FUNCTION "Get Station Selection Number" : Void   // FC16, SCL
{ S7_Optimized_Access := 'TRUE' }
VERSION : 0.1
   VAR_INPUT
      next : Bool;   // 'next' or 'prev'
      prev : Bool;
      stations : "Stations";
   END_VAR
   VAR_IN_OUT
      selStnNumber : Int;
   END_VAR
   VAR_TEMP
      i : Int;
      stnCount : Int;
      stnSelected : Bool;
   END_VAR
BEGIN
   REGION "COPY TO LOCAL"
       #stnCount := "stnCount";
   END_REGION

   REGION "INITIALIZE INDEX"
       #i := #selStnNumber;
   END_REGION

   REGION "PREVIOUS MODE"

       REGION "DECREMENT"
           IF #prev THEN
               #i -= 1;
           END_IF;
       END_REGION

       REGION "LOW LIMIT ROLLOVER"
           IF #i < 0 THEN
               #i := #stnCount;
           END_IF;
       END_REGION

   END_REGION

   REGION "NEXT MODE"

       REGION "INCREMENT"
           IF #next THEN
               #i += 1;
           END_IF;
       END_REGION

       REGION "HIGH LIMIT ROLLOVER"
           IF #i > #stnCount THEN
               #i := 0;
           END_IF;
       END_REGION

   END_REGION

   REGION "COPY TO LOCAL"
       #stnSelected := #stations.me[#i].settings.selected;
   END_REGION

   REGION "FIND NEXT SELECTED STATION"
       WHILE NOT #stnSelected DO

           REGION "PREVIOUS MODE"

               REGION "DECREMENT"
                   IF #prev THEN
                       #i -= 1;
                   END_IF;
               END_REGION

               REGION "LOW LIMIT ROLLOVER"
                   IF #i < 0 THEN
                       #i := #stnCount;
                   END_IF;
               END_REGION

           END_REGION

           REGION "NEXT MODE"

               REGION "INCREMENT"
                   IF #next THEN
                       #i += 1;
                   END_IF;
               END_REGION

               REGION "HIGH LIMIT ROLLOVER"
                   IF #i > #stnCount THEN
                       #i := 0;
                   END_IF;
               END_REGION

           END_REGION

           REGION "SAVE WHILE CONDITION"
               #stnSelected := #stations.me[#i].settings.selected;
           END_REGION

       END_WHILE;
   END_REGION

   REGION "RETURN VALUE"
       #selStnNumber := #i;
   END_REGION
END_FUNCTION

FUNCTION "Populate Button Details" : Void   // FC17, SCL
{ S7_Optimized_Access := 'TRUE' }
VERSION : 0.1
   VAR_INPUT
      selStnNumber : Int;
      stations : "Stations";
   END_VAR
   VAR_IN_OUT
      settings : "Settings";
   END_VAR
   VAR_TEMP
      btnCount : Int;
      i : Int;
      partNumber : WString;
      pBtn : Int;
      timerWS : WString;
   END_VAR
BEGIN
   REGION "COPY TO LOCAL"
       #btnCount := "ptsPerStn";
   END_REGION

   REGION "FOR EACH BUTTON"
       FOR #i := 0 TO #btnCount DO

           REGION "CALCULATE BUTTON POINTER"
               IF #i MOD 2 = 0 THEN
                   #pBtn := 7 - #i / 2;
               END_IF;
               IF #i MOD 2 <> 0 THEN
                   #pBtn := 3 - #i / 2;
               END_IF;
           END_REGION

           REGION "BUTTON LABEL"
               #settings.viewingStation.btns[#i].label.value := "Strip Sign"(INT_TO_WSTRING(#i + 1));
           END_REGION

           REGION "ALLOTTED TIME"
               #timerWS := "Real to WString Timer"(#stations.me[#selStnNumber].presetTime.allotted[#pBtn]);
               #settings.viewingStation.btns[#i].alloted.value := #timerWS;
           END_REGION

           REGION "CRITICAL TIME"
               #timerWS := "Real to WString Timer"(#stations.me[#selStnNumber].presetTime.critical[#pBtn]);
               #settings.viewingStation.btns[#i].critical.value := #timerWS;
           END_REGION

           REGION "PART NUMBER"
               #partNumber := #stations.me[#selStnNumber].partNumbers[#pBtn];
               #settings.viewingStation.btns[#i].partNumber.value := #partNumber;
           END_REGION

       END_FOR;
   END_REGION
END_FUNCTION

FUNCTION "Assign Station Parameters" : Void   // FC18, SCL
{ S7_Optimized_Access := 'TRUE' }
VERSION : 0.1
   VAR_IN_OUT
      settings : "Settings";
      stations : "Stations";
   END_VAR
   VAR_TEMP
      dzEntered : Bool;
      dzLabel : WString;
      i : Int;
      lineEntered : Bool;
      lineLabel : WString;
      stnCount : Int;
      stnSelected : Bool;
   END_VAR
BEGIN
   REGION "COPY TO LOCAL"    
       #dzEntered := #settings.viewingStation.dzData.inputFinished;
       #lineEntered := #settings.viewingStation.lineData.inputFinished;
       #stnCount := "stnCount";
   END_REGION

   REGION "ON PARAMETER ENTRY"
       IF #dzEntered OR #lineEntered THEN

           REGION "TURN OFF THE LIGHTS"
               #settings.viewingStation.dzData.inputFinished := FALSE;
               #settings.viewingStation.lineData.inputFinished := FALSE;
           END_REGION

           REGION "FOR EACH STATION"
               FOR #i := 0 TO #stnCount DO

                   REGION "COPY TO LOCAL"
                       #stnSelected := #stations.me[#i].settings.selected;
                   END_REGION

                   REGION "ON SELECTED STATION"
                       IF #stnSelected THEN

                           REGION "ON DROP ZONE INPUT"
                               IF #dzEntered THEN

                                   REGION "GET FROM HMI"
                                       #dzLabel := #settings.viewingStation.dzData.value;
                                   END_REGION

                                   REGION "WRITE TO STATION PARAMETER"
                                       #stations.me[#i].dropZone := WSTRING_TO_USINT(#dzLabel);
                                   END_REGION

                               END_IF;
                           END_REGION

                           REGION "ON LINE LABEL INPUT"
                               IF #lineEntered THEN

                                   REGION "GET FROM HMI"
                                       #lineLabel := #settings.viewingStation.lineData.value;
                                   END_REGION

                                   REGION "WRITE TO STATION PARAMETER"
                                       #stations.me[#i].line := #lineLabel;
                                   END_REGION

                               END_IF;
                           END_REGION

                       END_IF;
                   END_REGION

               END_FOR;
           END_REGION

       END_IF;
   END_REGION
END_FUNCTION

FUNCTION "Animate Button Details" : Void   // FC19, SCL
{ S7_Optimized_Access := 'TRUE' }
VERSION : 0.1
   VAR_INPUT
      stations : "Stations";
   END_VAR
   VAR_IN_OUT
      settings : "Settings";
   END_VAR
   VAR_TEMP
      animate : USInt;
      btnCount : Int;
      btnSelected : Bool;
      deselected : USInt;
      i : Int;
      invisible : USInt;
      pBtn : Int;
      selected : USInt;
      selStnCount : Int;
      selStnNumber : Int;
   END_VAR
BEGIN
   REGION "COPY TO LOCAL"
       #btnCount := "ptsPerStn";
       #deselected := "BgGray";
       #invisible := "invisible";
       #selected := "BgLTe";
       #selStnCount := #settings.#stations.selCount;
       #selStnNumber := #settings.stations.selNumber;
   END_REGION

   REGION "ENABLE"
       IF #selStnCount >= 1 THEN

           REGION "SHOW BUTTON DETAILS"
               #animate := #deselected;
           END_REGION

       END_IF;
   END_REGION

   REGION "DISABLE"
       IF #selStnCount = 0 THEN

           REGION "HIDE BUTTON DETAILS"
               #animate := #invisible;
           END_REGION

       END_IF;
   END_REGION

   REGION "APPLY ANIMATION"
       FOR #i := 0 TO #btnCount DO

           REGION "CALCULATE BUTTON POINTER"
               #pBtn := "Pointer Calc: Button Details"(#i);
           END_REGION

           REGION "WHILE Station SELECTED"
               IF #selStnCount <> 0 THEN

                   REGION "COPY TO LOCAL"
                       #btnSelected := #stations.me[#selStnNumber].settings.btnSelection[#pBtn];
                   END_REGION

                   REGION "ANIMATE BUTTON SELECTION

                       REGION "SELECTED"
                           IF #btnSelected THEN
                               #animate := #selected;
                           END_IF;
                       END_REGION

                       REGION "NOT SELECTED"
                           IF NOT #btnSelected THEN
                               #animate := #deselected;
                           END_IF;
                       END_REGION

                   END_REGION

               END_IF;
           END_REGION


           REGION "SEND TO HMI"
               #settings.viewingStation.btns[#i].label.animate := #animate;
               #settings.viewingStation.btns[#i].alloted.animate := #animate;
               #settings.viewingStation.btns[#i].critical.animate := #animate;
               #settings.viewingStation.btns[#i].partNumber.animate := #animate;
           END_REGION

       END_FOR;
   END_REGION
END_FUNCTION

FUNCTION "Populate Station Name" : WString   // FC20, SCL
{ S7_Optimized_Access := 'TRUE' }
VERSION : 0.1
   VAR_INPUT
      line : WString;
      dropZone : USInt;
   END_VAR
BEGIN
   #"Populate Station Name" := CONCAT_WSTRING(IN1 := #line,
                                              IN2 := wstring#' ',
                                              IN3 := "Strip Sign"(USINT_TO_WSTRING(#dropZone)));
END_FUNCTION

FUNCTION "Pointer Calc: Button Details" : Int   // FC21, SCL
{ S7_Optimized_Access := 'TRUE' }
VERSION : 0.1
   VAR_INPUT
      index : Int;
   END_VAR
   VAR_TEMP
      val : Int;
   END_VAR
BEGIN
   IF #index MOD 2 = 0 THEN
       #val := 7 - #index / 2;
   END_IF;

   IF #index MOD 2 <> 0 THEN
       #val := 3 - #index / 2;
   END_IF;

   #"Pointer Calc: Button Details" := #val;
END_FUNCTION

FUNCTION "Buffer Part Req Log Row: Generate" : "Part Req Log Row"   // FC22, SCL
{ S7_Optimized_Access := 'TRUE' }
VERSION : 0.1
   VAR_INPUT
      address : Int;
      "type" : Int;
   END_VAR
   VAR_TEMP
      retVal : Int;
   END_VAR
BEGIN
   REGION "ADDRESS"
       #"Buffer Part Req Log Row: Generate".address := #address;
   END_REGION

   REGION "REQUEST TYPE"
       #"Buffer Part Req Log Row: Generate".reqType := #type;
   END_REGION

   REGION "TIME STAMP"
       #retVal := RD_SYS_T(#"Buffer Part Req Log Row: Generate".timeStamp);
   END_REGION
END_FUNCTION

FUNCTION "Sim to Global" : Void   // FC23, SCL
{ S7_Optimized_Access := 'TRUE' }
VERSION : 0.1
   VAR_INPUT
      simStations : "Simulated Stations";
   END_VAR
   VAR_IN_OUT
      stations : "Stations";
   END_VAR
   VAR_TEMP
      btnCount : Int;
      firstStn : Int;
      i : Int;
      j : Int;
      pSim : Int;
      pStn : Int;
      simKP8Count : Int;
      stnCount : Int;
   END_VAR
BEGIN
   REGION "COPY TO LOCAL"
       #btnCount := "ptsPerStn";
       #firstStn := #simStations.firstStn;
       #simKP8Count := "simKP8Count";
       #stnCount := "stnCount";
   END_REGION

   REGION "FOR EACH STATION"
       FOR #i := 0 TO #simKP8Count DO

           REGION "CALCULATE POINTER"
               #pStn := #i + #firstStn;
               #pSim := #i;
           END_REGION

           REGION "UPPER LIMIT ROLL OVER"
               IF #pStn > #stnCount THEN
                   #pStn := #firstStn + #i - #stnCount - 1;
               END_IF;
           END_REGION

           REGION "COPY SIMULATED PRESSES"
               #stations.me[#pStn].kp8In := #simStations.me[#pSim].btn.actuate;
           END_REGION

       END_FOR;
   END_REGION
END_FUNCTION

FUNCTION "Pointer Calc: KP8 Labels" : Int   // FC25, SCL
{ S7_Optimized_Access := 'TRUE' }
VERSION : 0.1
   VAR_INPUT
      index : Int;
   END_VAR
   VAR_TEMP
      val : Int;
   END_VAR
BEGIN
   IF #index >= 4 THEN
       #val := 7 - (#index - 4) * 2;
   END_IF;

   IF #index <= 3 THEN
       #val := 8 - #index * 2;
   END_IF;

   #"Pointer Calc: KP8 Labels" := #val;
END_FUNCTION

FUNCTION "KP8 Color to Sim Animation" : USInt   // FC26, SCL
{ S7_Optimized_Access := 'TRUE' }
VERSION : 0.1
   VAR_INPUT
      kp8Color : DWord;
      btnNumber : Int;
   END_VAR
   VAR_TEMP
      animate : USInt;
      blue : USInt;
      colorDWord : DWord;
      colorInt : DInt;
      green : USInt;
      off : USInt;
      red : USInt;
      white : USInt;
      yellow : USInt;
   END_VAR
   VAR CONSTANT
      blueMask : DInt := 16#0000_0100;
      btnMask : DInt := 16#0101_0100;
      greenMask : DInt := 16#0001_0000;
      offMask : DInt := 16#0000_0000;
      redMask : DInt := 16#0100_0000;
      whiteMask : DInt := 16#0101_0100;
      yellowMask : DInt := 16#0101_0000;
   END_VAR
BEGIN
   REGION "COPY TO LOCAL"
       #blue := "BgLBl";
       #green := "BgLGr";
       #off := "BgGray";
       #red := "BgLRd";
       #white := "BgWh";
       #yellow := "BgLYe";
   END_REGION

   REGION "ISOLATE BUTTON COLOR"
       #colorDWord := SHR_DWORD(IN := #kp8Color,N := INT_TO_ULINT(#btnNumber));
       #colorDWord := #colorDWord AND #btnMask;
       #colorInt := DWORD_TO_DINT(#colorDWord);
   END_REGION

   REGION "DETERMINE ANIMATION"
       CASE #colorInt OF
           #blueMask:
               #animate := #blue;
           #greenMask:
               #animate := #green;
           #redMask:
               #animate := #red;
           #whiteMask:
               #animate := #white;
           #yellowMask:
               #animate := #yellow;
           ELSE
               #animate := #off;
       END_CASE;
   END_REGION

   REGION "RETURN VALUE"
       #"KP8 Color to Sim Animation" := #animate;
   END_REGION
END_FUNCTION

FUNCTION "Word Wrap" : WString   // FC28, SCL
{ S7_Optimized_Access := 'TRUE' }
VERSION : 0.1
   VAR_INPUT
      stringIn : WString;
      maxLength : Int;
   END_VAR
   VAR_TEMP
      length : Int;
      charBox : Array[0.."lStringLen"] of WChar;
      stringBox : Array[0.."lStringLen"] of WString["lStringLen"];
      count : UInt;
      status : Int;
      i : Int;
      pStringBox : Int;
      output : WString;
      savedOutput : WString;
      lineBox : Array[0..10] of WString["lStringLen"];
      pLineBox : Int;
      lengthTest : WString;
   END_VAR
   VAR CONSTANT
      space : WString := WSTRING#' ';
      blank : WString;
      lineBreak : WString := WSTRING#'$L';
   END_VAR
BEGIN
   #length := LEN(#stringIn);

   IF #length <= #maxLength THEN
       #output := #stringIn;
   END_IF;

   IF #length > #maxLength THEN

       Strg_TO_Chars(
                     Strg := #stringIn,
                     pChars := 0,
                     Cnt => #count,
                     Chars := #charBox
       );

       FOR #i := 0 TO "lStringLen" DO

           IF #charBox[#i] = #space THEN
               IF #charBox[#i + 1] = #space THEN
                   EXIT;
               END_IF;
           END_IF;

           IF #i = 0 THEN
               #stringBox[#pStringBox] := #charBox[#i];
           END_IF;

           IF #i >= 1 THEN
               #stringBox[#pStringBox] := CONCAT_WSTRING(IN1 := #stringBox[#pStringBox],
                                                         IN2 := #charBox[#i]);
           END_IF;

           IF #charBox[#i] = #space THEN
               #stringBox[#pStringBox] := "Trim"(#stringBox[#pStringBox]);
               #pStringBox := #pStringBox + 1;
           END_IF;

           IF #charBox[#i] = #lineBreak THEN
               #stringBox[#pStringBox] := LEFT(IN := #stringBox[#pStringBox],
                                               L := LEN(#stringBox[#pStringBox]) - 1);
               #pStringBox := #pStringBox + 1;
               #stringBox[#pStringBox] := #lineBreak;
               #pStringBox := #pStringBox + 1;
           END_IF;

       END_FOR;


       FOR #i := 0 TO "lStringLen" DO

           IF #stringBox[#i] = #blank THEN
               IF #stringBox[#i + 1] = #blank THEN
                   #lineBox[#pLineBox] := "Trim"(#lineBox[#pLineBox]);
                   EXIT;
               END_IF;
           END_IF;

           IF #stringBox[#i] = #lineBreak THEN
               #lineBox[#pLineBox] := "Trim"(#lineBox[#pLineBox]);
               #pLineBox := #pLineBox + 1;
               #lineBox[#pLineBox] := #lineBreak;
               #pLineBox := #pLineBox + 1;
           END_IF;


           IF #stringBox[#i] <> #lineBreak THEN

               IF #i = 0 THEN
                   #lengthTest := #stringBox[#i];
               END_IF;

               IF #i >= 1 THEN
                   #lengthTest := CONCAT_WSTRING(IN1 := #lineBox[#pLineBox],
                                                 IN2 := #space,
                                                 IN3 := #stringBox[#i]);
               END_IF;

               IF LEN(#lengthTest) <= #maxLength THEN
                   #lineBox[#pLineBox] := #lengthTest;
               END_IF;

               IF LEN(#lengthTest) > #maxLength THEN
                   #lineBox[#pLineBox] := "Trim"(#lineBox[#pLineBox]);
                   #lineBox[#pLineBox] := "Trim"(#lineBox[#pLineBox]);
                   #pLineBox := #pLineBox + 1;
                   #lineBox[#pLineBox] := #stringBox[#i];
               END_IF;
           END_IF;

       END_FOR;

       FOR #i := 0 TO 10 DO

           IF #lineBox[#i] = #space OR #lineBox[#i] = WString#'' THEN
               EXIT;
           END_IF;
           IF #i = 0 THEN
               #output := #lineBox[#i];
           END_IF;
           IF #i >= 1 THEN
               IF #lineBox[#i] = #lineBreak THEN
                   #output := #output;
               END_IF;
               IF #lineBox[#i] <> #lineBreak THEN
                   #output := CONCAT_WSTRING(IN1 := #output,
                                             IN2 := #lineBreak,
                                             IN3 := #lineBox[#i]);
               END_IF;
           END_IF;

       END_FOR;

       #output := "Trim"(#output);

   END_IF;

   #"Word Wrap" := #output;
END_FUNCTION

FUNCTION "Trim" : WString   // FC29, SCL
{ S7_Optimized_Access := 'TRUE' }
VERSION : 0.1
   VAR_INPUT
      stringIn : WString;
   END_VAR
   VAR_TEMP
      output : WString;
   END_VAR
   VAR CONSTANT
      space : WString := WSTRING#' ';
   END_VAR
BEGIN
   #output := #stringIn;
   IF LEFT(IN := #output, L := 1) = #space THEN
       #output := RIGHT(IN := #output, L := LEN(#output) - 1);
   END_IF;
   IF RIGHT(IN := #output, L := 1) = #space THEN
       #output := LEFT(IN := #output, L := LEN(#output) - 1);
   END_IF;
   #Trim := #output;
END_FUNCTION

FUNCTION "Recipe Select Button" : Void   // FC31, SCL
{ S7_Optimized_Access := 'TRUE' }
VERSION : 0.1
   VAR_INPUT
      visRows : Int;
      rowNum : Int;
      lib : "Menu: Library";
      actuate : Bool;
      maxRows : Int;
      btnNum : Int;
   END_VAR
   VAR_IN_OUT
      recipeSelectScreen : "HSS: Menu Selection Screen";
   END_VAR
   VAR_TEMP
      eval : "HSS: Menu Selection Screen";
      pRowVisLbl : Int;
      pRowInvisLbl : Int;
      pRowTxt : Int;
      pRecipeTxt : Int;
      maxLen : Int;
   END_VAR
BEGIN
   REGION "COPY TO LOCAL"
       #eval := #recipeSelectScreen;
   END_REGION


   REGION "NARROW"
       IF #maxRows > #visRows THEN
           #pRowVisLbl := #btnNum + #visRows;
           #pRowInvisLbl := #btnNum + (3 * #visRows);
           #maxLen := 22;
       END_IF;
   END_REGION


   REGION "WIDE"
       IF #maxRows <= #visRows THEN
           #pRowVisLbl := #btnNum + (3 * #visRows);
           #pRowInvisLbl := #btnNum + #visRows + 1;
           #maxLen := 28;
       END_IF;
   END_REGION


   REGION "ROW COUNT INDEPENDENT"
       #pRowTxt := (#btnNum * 2) + #visRows;
       #pRecipeTxt := #pRowTxt + 1;
   END_REGION


   REGION "DRAW"
       #eval.animate[#pRowVisLbl] := "BgGray";
       #eval.animate[#pRowInvisLbl] := "invisible";
       #eval.txt[#pRowTxt] := "Strip Sign"(DINT_TO_WSTRING(#rowNum));
       #eval.txt[#pRecipeTxt] := "Word Wrap"(stringIn := #lib.entry[#rowNum],
                                             maxLength := #maxLen);
   END_REGION

   REGION "ACTUATION ANIMATION"
       IF #actuate THEN
           #eval.animate[#pRowVisLbl] := "BgLTe";
       END_IF;
   END_REGION


   REGION "COPY TO GLOBAL"
       #recipeSelectScreen := #eval;
   END_REGION
END_FUNCTION

FUNCTION "Recipe Nav Button" : Void   // FC32, SCL
{ S7_Optimized_Access := 'TRUE' }
VERSION : 0.1
   VAR_INPUT
      visRows : Int;
      actuate : Bool;
      maxRows : Int;
      btnNum : Int;
   END_VAR
   VAR_IN_OUT
      recipeSelectScreen : "HSS: Menu Selection Screen";
   END_VAR
   VAR_TEMP
      eval : "HSS: Menu Selection Screen";
      color : Int;
   END_VAR
BEGIN
   REGION "COPY TO LOCAL"
       #eval := #recipeSelectScreen;
   END_REGION


   REGION "NARROW"
       IF #maxRows > #visRows THEN
           #color := "BgGray";
       END_IF;
   END_REGION


   REGION "WIDE"
       IF #maxRows <= #visRows THEN
           #color := "invisible";
       END_IF;
   END_REGION


   REGION "ROW COUNT INDEPENDENT"
       IF #actuate THEN
           #color := "BgLTe";
       END_IF;
   END_REGION


   REGION "DRAW"
       #eval.animate[#btnNum] := #color;
   END_REGION


   REGION "COPY TO GLOBAL"
       #recipeSelectScreen := #eval;
   END_REGION
END_FUNCTION

// ===== library types =====

TYPE "Table Row Data"
   STRUCT
      address : UInt;
      ordered : Bool;
      pbSelection : Struct
         actuate : Bool;
         animate : USInt;
      END_STRUCT;
      rtBackground : Struct
         animate : USInt;
      END_STRUCT;
      tfDropZone : Struct
         animate : USInt;
         value : WString[20];
      END_STRUCT;
      tfLine : Struct
         animate : USInt;
         value : WString[20];
      END_STRUCT;
      tfPartNumber : Struct
         animateDL : USInt;
         animateSL : USInt;
         value : WString[40];
      END_STRUCT;
      tfTime : Struct
         animate : USInt;
         value : WString[20];
      END_STRUCT;
   END_STRUCT;
END_TYPE

TYPE "Station Assignment: Button Details Data"
   STRUCT
      alloted : Struct
         animate : USInt;
         value : WString[10];
      END_STRUCT;
      critical : Struct
         animate : USInt;
         value : WString[10];
      END_STRUCT;
      label : Struct
         animate : USInt;
         value : WString[2];
      END_STRUCT;
      partNumber : Struct
         animate : USInt;
         value : WString[40];
      END_STRUCT;
      select : Struct
         actuate : Bool;
         animate : USInt;
      END_STRUCT;
   END_STRUCT;
END_TYPE

(* ===== HMI "HMI_RT_1" =====
system functions are stored by id; their names below are inferred from use
connection "HMI_Connection_2": ETHERNET, S7_1500_OMS

HMI tags "Default tag table"
   "Clock_Byte" : Byte = PLC Clock_Byte AT %MB0, 100 ms
   "HMI_screenNumber" : Int = PLC HMI.screenNumber AT %DB1.DBW0, 100 ms
   "HMI_barcode" : Barcode Screen = PLC HMI.barcode AT %DB1.DBW0, 100 ms
   "HMI_partCall_row{0}" : Table Row = PLC HMI.partCall.row[0], 100 ms
   "HMI_partCall_row{1}" : Table Row = PLC HMI.partCall.row[1], 100 ms
   "HMI_partCall_row{2}" : Table Row = PLC HMI.partCall.row[2], 100 ms
   "HMI_partCall_row{3}" : Table Row = PLC HMI.partCall.row[3], 100 ms
   "HMI_partCall_row{4}" : Table Row = PLC HMI.partCall.row[4], 100 ms
   "HMI_partCall_row{5}" : Table Row = PLC HMI.partCall.row[5], 100 ms
   "HMI_partCall_row{6}" : Table Row = PLC HMI.partCall.row[6], 100 ms
   "HMI_partCall_row{7}" : Table Row = PLC HMI.partCall.row[7], 100 ms
   "HMI_partCall_row{8}" : Table Row = PLC HMI.partCall.row[8], 100 ms
   "HMI_partCall_row{9}" : Table Row = PLC HMI.partCall.row[9], 100 ms
   "HMI_partCall_row{10}" : Table Row = PLC HMI.partCall.row[10], 100 ms
   "HMI_settings_stations_selectBtns{0}" : PB Data: Text Label = PLC HMI.settings.stations.selectBtns[0], 100 ms
   "HMI_settings_stations_selectBtns{1}" : PB Data: Text Label = PLC HMI.settings.stations.selectBtns[1], 100 ms
   "HMI_settings_stations_selectBtns{2}" : PB Data: Text Label = PLC HMI.settings.stations.selectBtns[2], 100 ms
   "HMI_settings_stations_selectBtns{3}" : PB Data: Text Label = PLC HMI.settings.stations.selectBtns[3], 100 ms
   "HMI_settings_stations_selectBtns{4}" : PB Data: Text Label = PLC HMI.settings.stations.selectBtns[4], 100 ms
   "HMI_settings_stations_selectBtns{5}" : PB Data: Text Label = PLC HMI.settings.stations.selectBtns[5], 100 ms
   "HMI_settings_stations_selectBtns{6}" : PB Data: Text Label = PLC HMI.settings.stations.selectBtns[6], 100 ms
   "HMI_settings_stations_selectBtns{7}" : PB Data: Text Label = PLC HMI.settings.stations.selectBtns[7], 100 ms
   "HMI_settings_stations_selectBtns{8}" : PB Data: Text Label = PLC HMI.settings.stations.selectBtns[8], 100 ms
   "HMI_settings_stations_selectBtns{9}" : PB Data: Text Label = PLC HMI.settings.stations.selectBtns[9], 100 ms
   "HMI_settings_stations_selectBtns{10}" : PB Data: Text Label = PLC HMI.settings.stations.selectBtns[10], 100 ms
   "HMI_settings_stations_selectBtns{11}" : PB Data: Text Label = PLC HMI.settings.stations.selectBtns[11], 100 ms
   "HMI_settings_kp8_buttons{0}" : PB Data: Text Label = PLC HMI.settings.kp8.buttons[0], 100 ms
   "HMI_settings_kp8_buttons{7}" : PB Data: Text Label = PLC HMI.settings.kp8.buttons[7], 100 ms
   "HMI_settings_kp8_buttons{3}" : PB Data: Text Label = PLC HMI.settings.kp8.buttons[3], 100 ms
   "HMI_settings_kp8_buttons{6}" : PB Data: Text Label = PLC HMI.settings.kp8.buttons[6], 100 ms
   "HMI_settings_kp8_buttons{2}" : PB Data: Text Label = PLC HMI.settings.kp8.buttons[2], 100 ms
   "HMI_settings_kp8_buttons{5}" : PB Data: Text Label = PLC HMI.settings.kp8.buttons[5], 100 ms
   "HMI_settings_kp8_buttons{1}" : PB Data: Text Label = PLC HMI.settings.kp8.buttons[1], 100 ms
   "HMI_settings_kp8_buttons{4}" : PB Data: Text Label = PLC HMI.settings.kp8.buttons[4], 100 ms
   "HMI_settings_stations_selCount" : Int = PLC HMI.settings.stations.selCount, 100 ms
   "HMI_settings_viewingStation_btns{0}" : Station Assignment: Button Details = PLC HMI.settings.viewingStation.btns[0], 100 ms
   "HMI_settings_viewingStation_btns{1}" : Station Assignment: Button Details = PLC HMI.settings.viewingStation.btns[1], 100 ms
   "HMI_settings_viewingStation_btns{2}" : Station Assignment: Button Details = PLC HMI.settings.viewingStation.btns[2], 100 ms
   "HMI_settings_viewingStation_btns{3}" : Station Assignment: Button Details = PLC HMI.settings.viewingStation.btns[3], 100 ms
   "HMI_settings_viewingStation_btns{4}" : Station Assignment: Button Details = PLC HMI.settings.viewingStation.btns[4], 100 ms
   "HMI_settings_viewingStation_btns{5}" : Station Assignment: Button Details = PLC HMI.settings.viewingStation.btns[5], 100 ms
   "HMI_settings_viewingStation_previous" : PB Data: Graphic/Text List = PLC HMI.settings.viewingStation.previous, 100 ms
   "HMI_settings_viewingStation_next" : PB Data: Graphic/Text List = PLC HMI.settings.viewingStation.next, 100 ms
   "HMI_settings_stations_selectAll" : PB Data: Text Label = PLC HMI.settings.stations.selectAll, 100 ms
   "HMI_settings_partNumber_assign" : PB Data: Text Label = PLC HMI.settings.partNumber.assign, 100 ms
   "HMI_settings_partNumber_ioField" : IO Field Data: Part Number = PLC HMI.settings.partNumber.ioField, 100 ms
   "HMI_settings_alotted_assign" : PB Data: Text Label = PLC HMI.settings.alotted.assign, 100 ms
   "HMI_settings_alotted_ioField" : IO Field Data: Timers = PLC HMI.settings.alotted.ioField, 100 ms
   "HMI_settings_critical_assign" : PB Data: Text Label = PLC HMI.settings.critical.assign, 100 ms
   "HMI_settings_critical_ioField" : IO Field Data: Timers = PLC HMI.settings.critical.ioField, 100 ms
   "HMI_settings_kp8_selectButtons" : PB Data: Text Label = PLC HMI.settings.kp8.selectButtons, 100 ms
   "HMI_settings_viewingStation_dzData" : Drop Zone Data = PLC HMI.settings.viewingStation.dzData, 100 ms
   "HMI_settings_viewingStation_lineData" : Line Label Data = PLC HMI.settings.viewingStation.lineData, 100 ms
   "HMI_settings_stations_prevGroup" : PB Data: Graphic/Text List = PLC HMI.settings.stations.prevGroup, 100 ms
   "HMI_settings_stations_nextGroup" : PB Data: Graphic/Text List = PLC HMI.settings.stations.nextGroup, 100 ms
   "HMI_settings_viewingStation_name" : WString[20] = PLC HMI.settings.viewingStation.name, 100 ms
   "HMI_tableNav_top" : PB Data: Graphic/Text List = PLC HMI.tableNav.top, 100 ms
   "HMI_tableNav_pageUp" : PB Data: Graphic/Text List = PLC HMI.tableNav.pageUp, 100 ms
   "HMI_tableNav_lineUp" : PB Data: Graphic/Text List = PLC HMI.tableNav.lineUp, 100 ms
   "HMI_tableNav_lineDown" : PB Data: Graphic/Text List = PLC HMI.tableNav.lineDown, 100 ms
   "HMI_tableNav_pageDown" : PB Data: Graphic/Text List = PLC HMI.tableNav.pageDown, 100 ms
   "HMI_tableNav_bottom" : PB Data: Graphic/Text List = PLC HMI.tableNav.bottom, 100 ms
   "HMI_simStations_stations{0}" : Station Sim Data = PLC HMI.simStations.me[0] AT %DB1.DBX0.0, 100 ms
   "HMI_simStations_me{1}" : Station Sim Data = PLC HMI.simStations.me[1], 100 ms
   "HMI_simStations_me{2}" : Station Sim Data = PLC HMI.simStations.me[2], 100 ms
   "HMI_simStations_me{3}" : Station Sim Data = PLC HMI.simStations.me[3], 100 ms
   "HMI_simStations_me{4}" : Station Sim Data = PLC HMI.simStations.me[4], 100 ms
   "HMI_simStations_me{5}" : Station Sim Data = PLC HMI.simStations.me[5], 100 ms
   "HMI_simStations_me{6}" : Station Sim Data = PLC HMI.simStations.me[6], 100 ms
   "HMI_simStations_me{7}" : Station Sim Data = PLC HMI.simStations.me[7], 100 ms
   "HMI_simStations_me{8}" : Station Sim Data = PLC HMI.simStations.me[8], 100 ms
   "HMI_simStations_me{9}" : Station Sim Data = PLC HMI.simStations.me[9], 100 ms
   "HMI_simStations_me{10}" : Station Sim Data = PLC HMI.simStations.me[10], 100 ms
   "HMI_simStations_me{11}" : Station Sim Data = PLC HMI.simStations.me[11], 100 ms
   "HMI_simStations_up" : PB Data: Graphic/Text List = PLC HMI.simStations.up, 100 ms
   "HMI_simStations_down" : PB Data: Graphic/Text List = PLC HMI.simStations.down, 100 ms
   "Log Flag" : Int = PLC "Log Buffer".logFlag AT %DB1.DBW0, 100 ms
      on ChangeValue: function_abcfba0d("Log Buffer_partReq_me{0}_address"); function_abcfba0d("Log Buffer_partReq_me{0}_timeStamp"); function_abcfba0d("Log Buffer_partReq_me{0}_reqType")
   "Log Buffer_partReq_me{0}_address" : Int = PLC "Log Buffer".partReq.me[0].address, 100 ms
   "Log Buffer_partReq_me{0}_timeStamp" : DTL = PLC "Log Buffer".partReq.me[0].timeStamp, 100 ms
   "Log Buffer_partReq_me{0}_reqType" : Int = PLC "Log Buffer".partReq.me[0].reqType, 100 ms
   "HMI_networkHealth_pnioDevices{1}" : PB Data: Text Label = PLC HMI.networkHealth.pnioDevices[1], 100 ms
   "HMI_networkHealth_pnioDevices{2}" : PB Data: Text Label = PLC HMI.networkHealth.pnioDevices[2], 1 s
   "HMI_networkHealth_pnioDevices{3}" : PB Data: Text Label = PLC HMI.networkHealth.pnioDevices[3], 1 s
   "HMI_networkHealth_pnioDevices{4}" : PB Data: Text Label = PLC HMI.networkHealth.pnioDevices[4], 1 s
   "HMI_networkHealth_pnioDevices{5}" : PB Data: Text Label = PLC HMI.networkHealth.pnioDevices[5], 1 s
   "HMI_networkHealth_pnioDevices{6}" : PB Data: Text Label = PLC HMI.networkHealth.pnioDevices[6], 1 s
   "HMI_networkHealth_pnioDevices{7}" : PB Data: Text Label = PLC HMI.networkHealth.pnioDevices[7], 1 s
   "HMI_networkHealth_pnioDevices{8}" : PB Data: Text Label = PLC HMI.networkHealth.pnioDevices[8], 1 s
   "HMI_networkHealth_pnioDevices{9}" : PB Data: Text Label = PLC HMI.networkHealth.pnioDevices[9], 1 s
   "HMI_networkHealth_pnioDevices{10}" : PB Data: Text Label = PLC HMI.networkHealth.pnioDevices[10], 1 s
   "HMI_networkHealth_pnioDevices{11}" : PB Data: Text Label = PLC HMI.networkHealth.pnioDevices[11], 1 s
   "HMI_networkHealth_pnioDevices{12}" : PB Data: Text Label = PLC HMI.networkHealth.pnioDevices[12], 1 s
   "HMI_networkHealth_pnioDevices{13}" : PB Data: Text Label = PLC HMI.networkHealth.pnioDevices[13], 1 s
   "HMI_networkHealth_pnioDevices{16}" : PB Data: Text Label = PLC HMI.networkHealth.pnioDevices[16], 1 s
   "HMI_networkHealth_pnioDevices{14}" : PB Data: Text Label = PLC HMI.networkHealth.pnioDevices[14], 1 s
   "HMI_networkHealth_pnioDevices{15}" : PB Data: Text Label = PLC HMI.networkHealth.pnioDevices[15], 1 s
   "HMI_networkHealth_pnioDevices{17}" : PB Data: Text Label = PLC HMI.networkHealth.pnioDevices[17], 1 s
   "HMI_networkHealth_pnioDevices{18}" : PB Data: Text Label = PLC HMI.networkHealth.pnioDevices[18], 1 s
   "HMI_networkHealth_pnioDevices{19}" : PB Data: Text Label = PLC HMI.networkHealth.pnioDevices[19], 1 s
   "HMI_networkHealth_pnioDevices{20}" : PB Data: Text Label = PLC HMI.networkHealth.pnioDevices[20], 1 s
   "HMI_networkHealth_pnioDevices{21}" : PB Data: Text Label = PLC HMI.networkHealth.pnioDevices[21], 1 s
   "HMI_networkHealth_pnioDevices{22}" : PB Data: Text Label = PLC HMI.networkHealth.pnioDevices[22], 1 s
   "HMI_networkHealth_pnioDevices{31}" : PB Data: Text Label = PLC HMI.networkHealth.pnioDevices[31], 1 s
   "HMI_networkHealth_pnioDevices{32}" : PB Data: Text Label = PLC HMI.networkHealth.pnioDevices[32], 1 s
   "HMI_networkHealth_pnioDevices{29}" : PB Data: Text Label = PLC HMI.networkHealth.pnioDevices[29], 1 s
   "HMI_networkHealth_pnioDevices{30}" : PB Data: Text Label = PLC HMI.networkHealth.pnioDevices[30], 1 s
   "HMI_networkHealth_pnioDevices{27}" : PB Data: Text Label = PLC HMI.networkHealth.pnioDevices[27], 1 s
   "HMI_networkHealth_pnioDevices{28}" : PB Data: Text Label = PLC HMI.networkHealth.pnioDevices[28], 1 s
   "HMI_networkHealth_pnioDevices{23}" : PB Data: Text Label = PLC HMI.networkHealth.pnioDevices[23], 1 s
   "HMI_networkHealth_pnioDevices{24}" : PB Data: Text Label = PLC HMI.networkHealth.pnioDevices[24], 1 s
   "HMI_networkHealth_pnioDevices{25}" : PB Data: Text Label = PLC HMI.networkHealth.pnioDevices[25], 1 s
   "HMI_networkHealth_pnioDevices{26}" : PB Data: Text Label = PLC HMI.networkHealth.pnioDevices[26], 1 s
   "HMI_networkHealth_pnioDevices{33}" : PB Data: Text Label = PLC HMI.networkHealth.pnioDevices[33], 1 s
   "HMI_networkHealth_pnioDevices{34}" : PB Data: Text Label = PLC HMI.networkHealth.pnioDevices[34], 1 s
   "HMI_networkHealth_pnioDevices{35}" : PB Data: Text Label = PLC HMI.networkHealth.pnioDevices[35], 1 s
   "HMI_networkHealth_pnioDevices{36}" : PB Data: Text Label = PLC HMI.networkHealth.pnioDevices[36], 1 s
   "HMI_networkHealth_pnioDevices{37}" : PB Data: Text Label = PLC HMI.networkHealth.pnioDevices[37], 1 s
   "HMI_networkHealth_pnioDevices{38}" : PB Data: Text Label = PLC HMI.networkHealth.pnioDevices[38], 1 s
   "HMI_networkHealth_pnioDevices{39}" : PB Data: Text Label = PLC HMI.networkHealth.pnioDevices[39], 1 s
   "HMI_networkHealth_pnioDevices{40}" : PB Data: Text Label = PLC HMI.networkHealth.pnioDevices[40], 1 s
   "HMI_networkHealth_pnioDevices{41}" : PB Data: Text Label = PLC HMI.networkHealth.pnioDevices[41], 1 s
   "HMI_networkHealth_pnioDevices{42}" : PB Data: Text Label = PLC HMI.networkHealth.pnioDevices[42], 1 s
   "HMI_networkHealth_pnioDevices{43}" : PB Data: Text Label = PLC HMI.networkHealth.pnioDevices[43], 1 s
   "HMI_networkHealth_pnioDevices{44}" : PB Data: Text Label = PLC HMI.networkHealth.pnioDevices[44], 1 s
   "HMI_networkHealth_pnioDevices{45}" : PB Data: Text Label = PLC HMI.networkHealth.pnioDevices[45], 1 s
   "HMI_networkHealth_pnioDevices{46}" : PB Data: Text Label = PLC HMI.networkHealth.pnioDevices[46], 1 s
   "HMI_networkHealth_pnioDevices{47}" : PB Data: Text Label = PLC HMI.networkHealth.pnioDevices[47], 1 s
   "HMI_networkHealth_pnioDevices{48}" : PB Data: Text Label = PLC HMI.networkHealth.pnioDevices[48], 1 s
   "HMI_networkHealth_et200spPopUp" : Station: ET200SP Comm Debug Data = PLC HMI.networkHealth.et200spPopUp, 1 s
   "HMI_networkHealth_kp8PopUp" : Station: KP8 Comm Debug Data = PLC HMI.networkHealth.kp8PopUp, 1 s
   "HMI_networkHealth_selectedDevice" : Int = PLC HMI.networkHealth.selectedDevice, 1 s
   "EMP IDB_stations_me{0}_partNumbers{0}" : WString[40] = PLC "EMP IDB".stations.me[0].partNumbers[0], 1 s
   "EMP IDB_stations_me{0}_partNumbers{1}" : WString[40] = PLC "EMP IDB".stations.me[0].partNumbers[1], 1 s
   "EMP IDB_stations_me{0}_partNumbers{2}" : WString[40] = PLC "EMP IDB".stations.me[0].partNumbers[2], 1 s
   "EMP IDB_stations_me{0}_partNumbers{3}" : WString[40] = PLC "EMP IDB".stations.me[0].partNumbers[3], 1 s
   "EMP IDB_stations_me{0}_partNumbers{4}" : WString[40] = PLC "EMP IDB".stations.me[0].partNumbers[4], 1 s
   "EMP IDB_stations_me{0}_partNumbers{5}" : WString[40] = PLC "EMP IDB".stations.me[0].partNumbers[5], 1 s
   "EMP IDB_stations_me{0}_partNumbers{6}" : WString[40] = PLC "EMP IDB".stations.me[0].partNumbers[6], 1 s
   "EMP IDB_stations_me{0}_partNumbers{7}" : WString[40] = PLC "EMP IDB".stations.me[0].partNumbers[7], 1 s
   "EMP IDB_stations_me{1}_partNumbers{0}" : WString[40] = PLC "EMP IDB".stations.me[1].partNumbers[0], 1 s
   "EMP IDB_stations_me{1}_partNumbers{1}" : WString[40] = PLC "EMP IDB".stations.me[1].partNumbers[1], 1 s
   "EMP IDB_stations_me{1}_partNumbers{2}" : WString[40] = PLC "EMP IDB".stations.me[1].partNumbers[2], 1 s
   "EMP IDB_stations_me{1}_partNumbers{3}" : WString[40] = PLC "EMP IDB".stations.me[1].partNumbers[3], 1 s
   "EMP IDB_stations_me{1}_partNumbers{4}" : WString[40] = PLC "EMP IDB".stations.me[1].partNumbers[4], 1 s
   "EMP IDB_stations_me{1}_partNumbers{5}" : WString[40] = PLC "EMP IDB".stations.me[1].partNumbers[5], 1 s
   "EMP IDB_stations_me{1}_partNumbers{6}" : WString[40] = PLC "EMP IDB".stations.me[1].partNumbers[6], 1 s
   "EMP IDB_stations_me{1}_partNumbers{7}" : WString[40] = PLC "EMP IDB".stations.me[1].partNumbers[7], 1 s
   "EMP IDB_stations_me{2}_partNumbers{0}" : WString[40] = PLC "EMP IDB".stations.me[2].partNumbers[0], 1 s
   "EMP IDB_stations_me{2}_partNumbers{1}" : WString[40] = PLC "EMP IDB".stations.me[2].partNumbers[1], 1 s
   "EMP IDB_stations_me{2}_partNumbers{2}" : WString[40] = PLC "EMP IDB".stations.me[2].partNumbers[2], 1 s
   "EMP IDB_stations_me{2}_partNumbers{3}" : WString[40] = PLC "EMP IDB".stations.me[2].partNumbers[3], 1 s
   "EMP IDB_stations_me{2}_partNumbers{4}" : WString[40] = PLC "EMP IDB".stations.me[2].partNumbers[4], 1 s
   "EMP IDB_stations_me{2}_partNumbers{5}" : WString[40] = PLC "EMP IDB".stations.me[2].partNumbers[5], 1 s
   "EMP IDB_stations_me{2}_partNumbers{6}" : WString[40] = PLC "EMP IDB".stations.me[2].partNumbers[6], 1 s
   "EMP IDB_stations_me{2}_partNumbers{7}" : WString[40] = PLC "EMP IDB".stations.me[2].partNumbers[7], 1 s
   "EMP IDB_stations_me{3}_partOrdered{0}" : Bool = PLC "EMP IDB".stations.me[3].partOrdered[0], 1 s
   "EMP IDB_stations_me{3}_partOrdered{1}" : Bool = PLC "EMP IDB".stations.me[3].partOrdered[1], 1 s
   "EMP IDB_stations_me{3}_partOrdered{2}" : Bool = PLC "EMP IDB".stations.me[3].partOrdered[2], 1 s
   "EMP IDB_stations_me{3}_partOrdered{3}" : Bool = PLC "EMP IDB".stations.me[3].partOrdered[3], 1 s
   "EMP IDB_stations_me{3}_partOrdered{4}" : Bool = PLC "EMP IDB".stations.me[3].partOrdered[4], 1 s
   "EMP IDB_stations_me{3}_partOrdered{5}" : Bool = PLC "EMP IDB".stations.me[3].partOrdered[5], 1 s
   "EMP IDB_stations_me{3}_partOrdered{6}" : Bool = PLC "EMP IDB".stations.me[3].partOrdered[6], 1 s
   "EMP IDB_stations_me{3}_partOrdered{7}" : Bool = PLC "EMP IDB".stations.me[3].partOrdered[7], 1 s
   "EMP IDB_stations_me{4}_partNumbers{0}" : WString[40] = PLC "EMP IDB".stations.me[4].partNumbers[0], 1 s
   "EMP IDB_stations_me{4}_partNumbers{1}" : WString[40] = PLC "EMP IDB".stations.me[4].partNumbers[1], 1 s
   "EMP IDB_stations_me{4}_partNumbers{2}" : WString[40] = PLC "EMP IDB".stations.me[4].partNumbers[2], 1 s
   "EMP IDB_stations_me{4}_partNumbers{3}" : WString[40] = PLC "EMP IDB".stations.me[4].partNumbers[3], 1 s
   "EMP IDB_stations_me{4}_partNumbers{4}" : WString[40] = PLC "EMP IDB".stations.me[4].partNumbers[4], 1 s
   "EMP IDB_stations_me{4}_partNumbers{5}" : WString[40] = PLC "EMP IDB".stations.me[4].partNumbers[5], 1 s
   "EMP IDB_stations_me{4}_partNumbers{6}" : WString[40] = PLC "EMP IDB".stations.me[4].partNumbers[6], 1 s
   "EMP IDB_stations_me{4}_partNumbers{7}" : WString[40] = PLC "EMP IDB".stations.me[4].partNumbers[7], 1 s
   "EMP IDB_stations_me{5}_partNumbers{0}" : WString[40] = PLC "EMP IDB".stations.me[5].partNumbers[0], 1 s
   "EMP IDB_stations_me{5}_partNumbers{1}" : WString[40] = PLC "EMP IDB".stations.me[5].partNumbers[1], 1 s
   "EMP IDB_stations_me{5}_partNumbers{2}" : WString[40] = PLC "EMP IDB".stations.me[5].partNumbers[2], 1 s
   "EMP IDB_stations_me{5}_partNumbers{3}" : WString[40] = PLC "EMP IDB".stations.me[5].partNumbers[3], 1 s
   "EMP IDB_stations_me{5}_partNumbers{4}" : WString[40] = PLC "EMP IDB".stations.me[5].partNumbers[4], 1 s
   "EMP IDB_stations_me{5}_partNumbers{5}" : WString[40] = PLC "EMP IDB".stations.me[5].partNumbers[5], 1 s
   "EMP IDB_stations_me{5}_partNumbers{6}" : WString[40] = PLC "EMP IDB".stations.me[5].partNumbers[6], 1 s
   "EMP IDB_stations_me{5}_partNumbers{7}" : WString[40] = PLC "EMP IDB".stations.me[5].partNumbers[7], 1 s
   "EMP IDB_stations_me{6}_partNumbers{0}" : WString[40] = PLC "EMP IDB".stations.me[6].partNumbers[0], 1 s
   "EMP IDB_stations_me{6}_partNumbers{1}" : WString[40] = PLC "EMP IDB".stations.me[6].partNumbers[1], 1 s
   "EMP IDB_stations_me{6}_partNumbers{2}" : WString[40] = PLC "EMP IDB".stations.me[6].partNumbers[2], 1 s
   "EMP IDB_stations_me{6}_partNumbers{3}" : WString[40] = PLC "EMP IDB".stations.me[6].partNumbers[3], 1 s
   "EMP IDB_stations_me{6}_partNumbers{4}" : WString[40] = PLC "EMP IDB".stations.me[6].partNumbers[4], 1 s
   "EMP IDB_stations_me{6}_partNumbers{5}" : WString[40] = PLC "EMP IDB".stations.me[6].partNumbers[5], 1 s
   "EMP IDB_stations_me{6}_partNumbers{6}" : WString[40] = PLC "EMP IDB".stations.me[6].partNumbers[6], 1 s
   "EMP IDB_stations_me{6}_partNumbers{7}" : WString[40] = PLC "EMP IDB".stations.me[6].partNumbers[7], 1 s
   "EMP IDB_stations_me{7}_partNumbers{0}" : WString[40] = PLC "EMP IDB".stations.me[7].partNumbers[0], 1 s
   "EMP IDB_stations_me{7}_partNumbers{1}" : WString[40] = PLC "EMP IDB".stations.me[7].partNumbers[1], 1 s
   "EMP IDB_stations_me{7}_partNumbers{2}" : WString[40] = PLC "EMP IDB".stations.me[7].partNumbers[2], 1 s
   "EMP IDB_stations_me{7}_partNumbers{3}" : WString[40] = PLC "EMP IDB".stations.me[7].partNumbers[3], 1 s
   "EMP IDB_stations_me{7}_partNumbers{4}" : WString[40] = PLC "EMP IDB".stations.me[7].partNumbers[4], 1 s
   "EMP IDB_stations_me{7}_partNumbers{5}" : WString[40] = PLC "EMP IDB".stations.me[7].partNumbers[5], 1 s
   "EMP IDB_stations_me{7}_partNumbers{6}" : WString[40] = PLC "EMP IDB".stations.me[7].partNumbers[6], 1 s
   "EMP IDB_stations_me{7}_partNumbers{7}" : WString[40] = PLC "EMP IDB".stations.me[7].partNumbers[7], 1 s
   "EMP IDB_stations_me{8}_partNumbers{0}" : WString[40] = PLC "EMP IDB".stations.me[8].partNumbers[0], 1 s
   "EMP IDB_stations_me{8}_partNumbers{1}" : WString[40] = PLC "EMP IDB".stations.me[8].partNumbers[1], 1 s
   "EMP IDB_stations_me{8}_partNumbers{2}" : WString[40] = PLC "EMP IDB".stations.me[8].partNumbers[2], 1 s
   "EMP IDB_stations_me{8}_partNumbers{3}" : WString[40] = PLC "EMP IDB".stations.me[8].partNumbers[3], 1 s
   "EMP IDB_stations_me{8}_partNumbers{4}" : WString[40] = PLC "EMP IDB".stations.me[8].partNumbers[4], 1 s
   "EMP IDB_stations_me{8}_partNumbers{5}" : WString[40] = PLC "EMP IDB".stations.me[8].partNumbers[5], 1 s
   "EMP IDB_stations_me{8}_partNumbers{6}" : WString[40] = PLC "EMP IDB".stations.me[8].partNumbers[6], 1 s
   "EMP IDB_stations_me{8}_partNumbers{7}" : WString[40] = PLC "EMP IDB".stations.me[8].partNumbers[7], 1 s
   "EMP IDB_stations_me{9}_partNumbers{0}" : WString[40] = PLC "EMP IDB".stations.me[9].partNumbers[0], 1 s
   "EMP IDB_stations_me{9}_partNumbers{1}" : WString[40] = PLC "EMP IDB".stations.me[9].partNumbers[1], 1 s
   "EMP IDB_stations_me{9}_partNumbers{2}" : WString[40] = PLC "EMP IDB".stations.me[9].partNumbers[2], 1 s
   "EMP IDB_stations_me{9}_partNumbers{3}" : WString[40] = PLC "EMP IDB".stations.me[9].partNumbers[3], 1 s
   "EMP IDB_stations_me{9}_partNumbers{4}" : WString[40] = PLC "EMP IDB".stations.me[9].partNumbers[4], 1 s
   "EMP IDB_stations_me{9}_partNumbers{5}" : WString[40] = PLC "EMP IDB".stations.me[9].partNumbers[5], 1 s
   "EMP IDB_stations_me{9}_partNumbers{6}" : WString[40] = PLC "EMP IDB".stations.me[9].partNumbers[6], 1 s
   "EMP IDB_stations_me{9}_partNumbers{7}" : WString[40] = PLC "EMP IDB".stations.me[9].partNumbers[7], 1 s
   "EMP IDB_stations_me{10}_partNumbers{0}" : WString[40] = PLC "EMP IDB".stations.me[10].partNumbers[0], 1 s
   "EMP IDB_stations_me{10}_partNumbers{1}" : WString[40] = PLC "EMP IDB".stations.me[10].partNumbers[1], 1 s
   "EMP IDB_stations_me{10}_partNumbers{2}" : WString[40] = PLC "EMP IDB".stations.me[10].partNumbers[2], 1 s
   "EMP IDB_stations_me{10}_partNumbers{3}" : WString[40] = PLC "EMP IDB".stations.me[10].partNumbers[3], 1 s
   "EMP IDB_stations_me{10}_partNumbers{4}" : WString[40] = PLC "EMP IDB".stations.me[10].partNumbers[4], 1 s
   "EMP IDB_stations_me{10}_partNumbers{5}" : WString[40] = PLC "EMP IDB".stations.me[10].partNumbers[5], 1 s
   "EMP IDB_stations_me{10}_partNumbers{6}" : WString[40] = PLC "EMP IDB".stations.me[10].partNumbers[6], 1 s
   "EMP IDB_stations_me{10}_partNumbers{7}" : WString[40] = PLC "EMP IDB".stations.me[10].partNumbers[7], 1 s
   "EMP IDB_stations_me{11}_partNumbers{0}" : WString[40] = PLC "EMP IDB".stations.me[11].partNumbers[0], 1 s
   "EMP IDB_stations_me{11}_partNumbers{1}" : WString[40] = PLC "EMP IDB".stations.me[11].partNumbers[1], 1 s
   "EMP IDB_stations_me{11}_partNumbers{2}" : WString[40] = PLC "EMP IDB".stations.me[11].partNumbers[2], 1 s
   "EMP IDB_stations_me{11}_partNumbers{3}" : WString[40] = PLC "EMP IDB".stations.me[11].partNumbers[3], 1 s
   "EMP IDB_stations_me{11}_partNumbers{4}" : WString[40] = PLC "EMP IDB".stations.me[11].partNumbers[4], 1 s
   "EMP IDB_stations_me{11}_partNumbers{5}" : WString[40] = PLC "EMP IDB".stations.me[11].partNumbers[5], 1 s
   "EMP IDB_stations_me{11}_partNumbers{6}" : WString[40] = PLC "EMP IDB".stations.me[11].partNumbers[6], 1 s
   "EMP IDB_stations_me{11}_partNumbers{7}" : WString[40] = PLC "EMP IDB".stations.me[11].partNumbers[7], 1 s
   "EMP IDB_stations_me{12}_partNumbers{0}" : WString[40] = PLC "EMP IDB".stations.me[12].partNumbers[0], 1 s
   "EMP IDB_stations_me{12}_partNumbers{1}" : WString[40] = PLC "EMP IDB".stations.me[12].partNumbers[1], 1 s
   "EMP IDB_stations_me{12}_partNumbers{2}" : WString[40] = PLC "EMP IDB".stations.me[12].partNumbers[2], 1 s
   "EMP IDB_stations_me{12}_partNumbers{3}" : WString[40] = PLC "EMP IDB".stations.me[12].partNumbers[3], 1 s
   "EMP IDB_stations_me{12}_partNumbers{4}" : WString[40] = PLC "EMP IDB".stations.me[12].partNumbers[4], 1 s
   "EMP IDB_stations_me{12}_partNumbers{5}" : WString[40] = PLC "EMP IDB".stations.me[12].partNumbers[5], 1 s
   "EMP IDB_stations_me{12}_partNumbers{6}" : WString[40] = PLC "EMP IDB".stations.me[12].partNumbers[6], 1 s
   "EMP IDB_stations_me{12}_partNumbers{7}" : WString[40] = PLC "EMP IDB".stations.me[12].partNumbers[7], 1 s
   "EMP IDB_stations_me{13}_partNumbers{0}" : WString[40] = PLC "EMP IDB".stations.me[13].partNumbers[0], 1 s
   "EMP IDB_stations_me{13}_partNumbers{1}" : WString[40] = PLC "EMP IDB".stations.me[13].partNumbers[1], 1 s
   "EMP IDB_stations_me{13}_partNumbers{2}" : WString[40] = PLC "EMP IDB".stations.me[13].partNumbers[2], 1 s
   "EMP IDB_stations_me{13}_partNumbers{3}" : WString[40] = PLC "EMP IDB".stations.me[13].partNumbers[3], 1 s
   "EMP IDB_stations_me{13}_partNumbers{4}" : WString[40] = PLC "EMP IDB".stations.me[13].partNumbers[4], 1 s
   "EMP IDB_stations_me{13}_partNumbers{5}" : WString[40] = PLC "EMP IDB".stations.me[13].partNumbers[5], 1 s
   "EMP IDB_stations_me{13}_partNumbers{6}" : WString[40] = PLC "EMP IDB".stations.me[13].partNumbers[6], 1 s
   "EMP IDB_stations_me{13}_partNumbers{7}" : WString[40] = PLC "EMP IDB".stations.me[13].partNumbers[7], 1 s
   "EMP IDB_stations_me{14}_partNumbers{0}" : WString[40] = PLC "EMP IDB".stations.me[14].partNumbers[0], 1 s
   "EMP IDB_stations_me{14}_partNumbers{1}" : WString[40] = PLC "EMP IDB".stations.me[14].partNumbers[1], 1 s
   "EMP IDB_stations_me{14}_partNumbers{2}" : WString[40] = PLC "EMP IDB".stations.me[14].partNumbers[2], 1 s
   "EMP IDB_stations_me{14}_partNumbers{3}" : WString[40] = PLC "EMP IDB".stations.me[14].partNumbers[3], 1 s
   "EMP IDB_stations_me{14}_partNumbers{4}" : WString[40] = PLC "EMP IDB".stations.me[14].partNumbers[4], 1 s
   "EMP IDB_stations_me{14}_partNumbers{5}" : WString[40] = PLC "EMP IDB".stations.me[14].partNumbers[5], 1 s
   "EMP IDB_stations_me{14}_partNumbers{6}" : WString[40] = PLC "EMP IDB".stations.me[14].partNumbers[6], 1 s
   "EMP IDB_stations_me{14}_partNumbers{7}" : WString[40] = PLC "EMP IDB".stations.me[14].partNumbers[7], 1 s
   "EMP IDB_stations_me{15}_partNumbers{0}" : WString[40] = PLC "EMP IDB".stations.me[15].partNumbers[0], 1 s
   "EMP IDB_stations_me{15}_partNumbers{1}" : WString[40] = PLC "EMP IDB".stations.me[15].partNumbers[1], 1 s
   "EMP IDB_stations_me{15}_partNumbers{2}" : WString[40] = PLC "EMP IDB".stations.me[15].partNumbers[2], 1 s
   "EMP IDB_stations_me{15}_partNumbers{3}" : WString[40] = PLC "EMP IDB".stations.me[15].partNumbers[3], 1 s
   "EMP IDB_stations_me{15}_partNumbers{4}" : WString[40] = PLC "EMP IDB".stations.me[15].partNumbers[4], 1 s
   "EMP IDB_stations_me{15}_partNumbers{5}" : WString[40] = PLC "EMP IDB".stations.me[15].partNumbers[5], 1 s
   "EMP IDB_stations_me{15}_partNumbers{6}" : WString[40] = PLC "EMP IDB".stations.me[15].partNumbers[6], 1 s
   "EMP IDB_stations_me{15}_partNumbers{7}" : WString[40] = PLC "EMP IDB".stations.me[15].partNumbers[7], 1 s
   "EMP IDB_stations_me{16}_partNumbers{0}" : WString[40] = PLC "EMP IDB".stations.me[16].partNumbers[0], 1 s
   "EMP IDB_stations_me{16}_partNumbers{1}" : WString[40] = PLC "EMP IDB".stations.me[16].partNumbers[1], 1 s